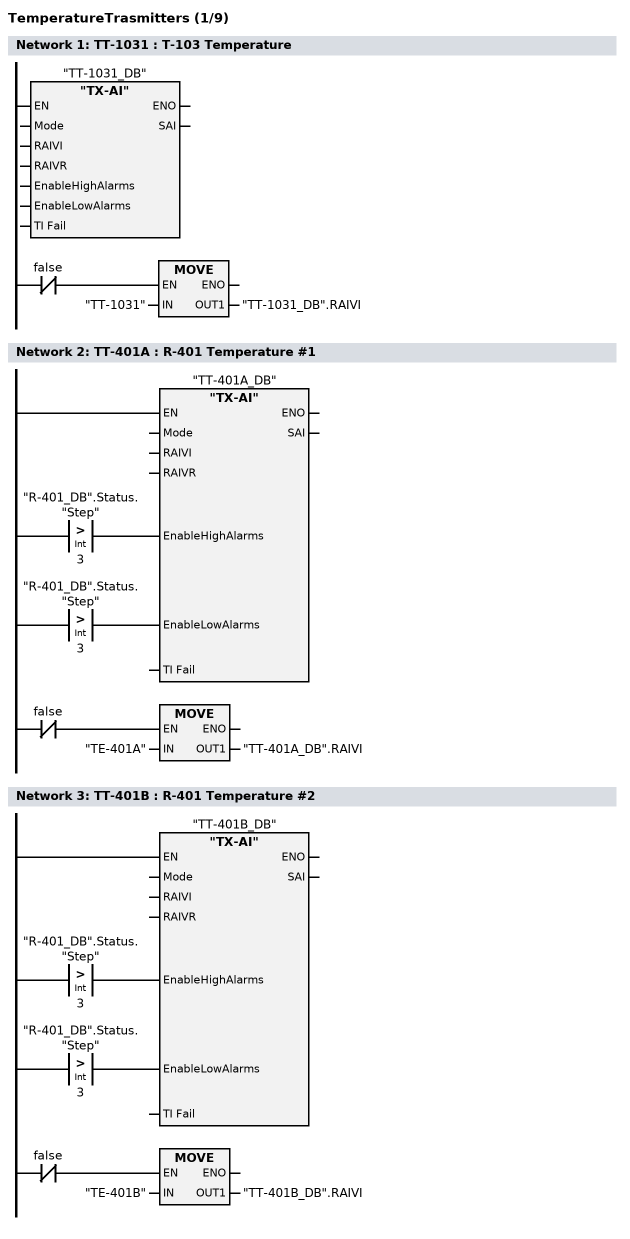
   RUNG wire#powerrail
      "TT-1031_DB"(Mode :=, RAIVI :=, RAIVR :=, EnableHighAlarms :=, EnableLowAlarms :=, "TI Fail" :=, SAI =>)
   END_RUNG
   RUNG wire#powerrail
      I_Contact( false )
      { S7_GenerateENO := "TRUE" } Move(in := "TT-1031", out1 => "TT-1031_DB".RAIVI)
   END_RUNG
   // the same network as SCL:
   "TT-1031_DB"();   // "TX-AI"
   IF NOT false THEN "TT-1031_DB".RAIVI := "TT-1031"; END_IF;
END_REGION

REGION Network 2: TT-401A : R-401 Temperature #1
   RUNG wire#powerrail
      "TT-401A_DB"(EnableHighAlarms := wire#w1, EnableLowAlarms := wire#w2, Mode :=, RAIVI :=, RAIVR :=, "TI Fail" :=, SAI =>)
   END_RUNG
   RUNG wire#powerrail
      { S7_Templates := "SrcType := Int" } GT_Contact(in1 := "R-401_DB".Status."Step", in2 := 3)
   END_RUNG wire#w1
   RUNG wire#powerrail
      { S7_Templates := "SrcType := Int" } GT_Contact(in1 := "R-401_DB".Status."Step", in2 := 3)
   END_RUNG wire#w2
   RUNG wire#powerrail
      I_Contact( false )
      { S7_GenerateENO := "TRUE" } Move(in := "TE-401A", out1 => "TT-401A_DB".RAIVI)
   END_RUNG
   // the same network as SCL:
   "TT-401A_DB"(EnableHighAlarms := "R-401_DB".Status."Step" > 3,   // "TX-AI"
                EnableLowAlarms := "R-401_DB".Status."Step" > 3);
   IF NOT false THEN "TT-401A_DB".RAIVI := "TE-401A"; END_IF;
END_REGION

REGION Network 3: TT-401B : R-401 Temperature #2
   RUNG wire#powerrail
      "TT-401B_DB"(EnableHighAlarms := wire#w1, EnableLowAlarms := wire#w2, Mode :=, RAIVI :=, RAIVR :=, "TI Fail" :=, SAI =>)
   END_RUNG
   RUNG wire#powerrail
      { S7_Templates := "SrcType := Int" } GT_Contact(in1 := "R-401_DB".Status."Step", in2 := 3)
   END_RUNG wire#w1
   RUNG wire#powerrail
      { S7_Templates := "SrcType := Int" } GT_Contact(in1 := "R-401_DB".Status."Step", in2 := 3)
   END_RUNG wire#w2
   RUNG wire#powerrail
      I_Contact( false )
      { S7_GenerateENO := "TRUE" } Move(in := "TE-401B", out1 => "TT-401B_DB".RAIVI)
   END_RUNG
   // the same network as SCL:
   "TT-401B_DB"(EnableHighAlarms := "R-401_DB".Status."Step" > 3,   // "TX-AI"
                EnableLowAlarms := "R-401_DB".Status."Step" > 3);
   IF NOT false THEN "TT-401B_DB".RAIVI := "TE-401B"; END_IF;
END_REGION

REGION Network 4: TT-401C : R-401 Temperature #3
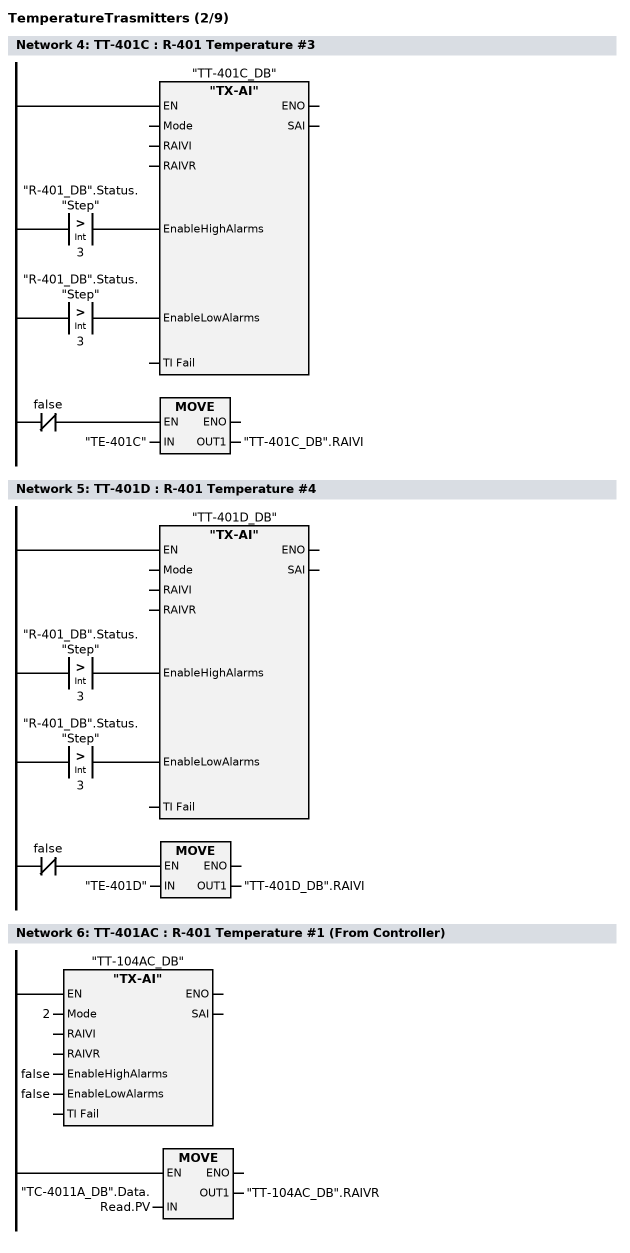
   RUNG wire#powerrail
      "TT-401C_DB"(EnableHighAlarms := wire#w1, EnableLowAlarms := wire#w2, Mode :=, RAIVI :=, RAIVR :=, "TI Fail" :=, SAI =>)
   END_RUNG
   RUNG wire#powerrail
      { S7_Templates := "SrcType := Int" } GT_Contact(in1 := "R-401_DB".Status."Step", in2 := 3)
   END_RUNG wire#w1
   RUNG wire#powerrail
      { S7_Templates := "SrcType := Int" } GT_Contact(in1 := "R-401_DB".Status."Step", in2 := 3)
   END_RUNG wire#w2
   RUNG wire#powerrail
      I_Contact( false )
      { S7_GenerateENO := "TRUE" } Move(in := "TE-401C", out1 => "TT-401C_DB".RAIVI)
   END_RUNG
   // the same network as SCL:
   "TT-401C_DB"(EnableHighAlarms := "R-401_DB".Status."Step" > 3,   // "TX-AI"
                EnableLowAlarms := "R-401_DB".Status."Step" > 3);
   IF NOT false THEN "TT-401C_DB".RAIVI := "TE-401C"; END_IF;
END_REGION

REGION Network 5: TT-401D : R-401 Temperature #4
   RUNG wire#powerrail
      "TT-401D_DB"(EnableHighAlarms := wire#w1, EnableLowAlarms := wire#w2, Mode :=, RAIVI :=, RAIVR :=, "TI Fail" :=, SAI =>)
   END_RUNG
   RUNG wire#powerrail
      { S7_Templates := "SrcType := Int" } GT_Contact(in1 := "R-401_DB".Status."Step", in2 := 3)
   END_RUNG wire#w1
   RUNG wire#powerrail
      { S7_Templates := "SrcType := Int" } GT_Contact(in1 := "R-401_DB".Status."Step", in2 := 3)
   END_RUNG wire#w2
   RUNG wire#powerrail
      I_Contact( false )
      { S7_GenerateENO := "TRUE" } Move(in := "TE-401D", out1 => "TT-401D_DB".RAIVI)
   END_RUNG
   // the same network as SCL:
   "TT-401D_DB"(EnableHighAlarms := "R-401_DB".Status."Step" > 3,   // "TX-AI"
                EnableLowAlarms := "R-401_DB".Status."Step" > 3);
   IF NOT false THEN "TT-401D_DB".RAIVI := "TE-401D"; END_IF;
END_REGION

REGION Network 6: TT-401AC : R-401 Temperature #1 (From Controller)
   RUNG wire#powerrail
      "TT-104AC_DB"(Mode := 2, RAIVI :=, RAIVR :=, EnableHighAlarms := false, EnableLowAlarms := false, "TI Fail" :=, SAI =>)
   END_RUNG
   RUNG wire#powerrail
      { S7_GenerateENO := "TRUE" } Move(in := "TC-4011A_DB".Data.Read.PV, out1 => "TT-104AC_DB".RAIVR)
   END_RUNG
   // the same network as SCL:
   "TT-104AC_DB"(Mode := 2, EnableHighAlarms := false, EnableLowAlarms := false);   // "TX-AI"
   "TT-104AC_DB".RAIVR := "TC-4011A_DB".Data.Read.PV;
END_REGION

REGION Network 7: TT-401BC : R-401 Temperature #2 (From Controller)
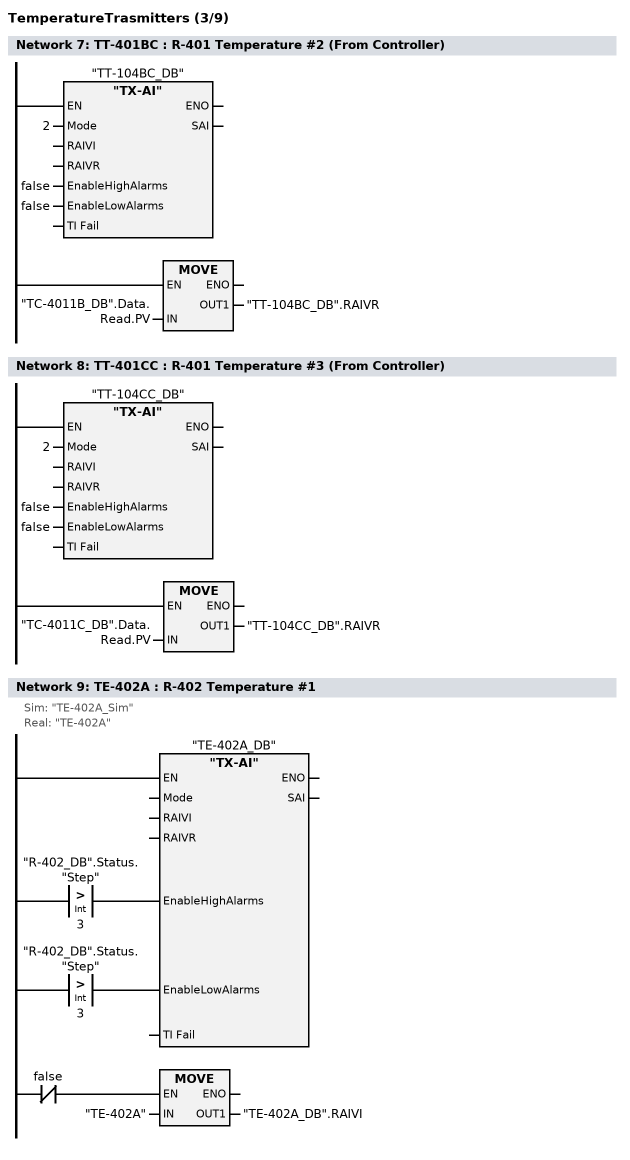
   RUNG wire#powerrail
      "TT-104BC_DB"(Mode := 2, RAIVI :=, RAIVR :=, EnableHighAlarms := false, EnableLowAlarms := false, "TI Fail" :=, SAI =>)
   END_RUNG
   RUNG wire#powerrail
      { S7_GenerateENO := "TRUE" } Move(in := "TC-4011B_DB".Data.Read.PV, out1 => "TT-104BC_DB".RAIVR)
   END_RUNG
   // the same network as SCL:
   "TT-104BC_DB"(Mode := 2, EnableHighAlarms := false, EnableLowAlarms := false);   // "TX-AI"
   "TT-104BC_DB".RAIVR := "TC-4011B_DB".Data.Read.PV;
END_REGION

REGION Network 8: TT-401CC : R-401 Temperature #3 (From Controller)
   RUNG wire#powerrail
      "TT-104CC_DB"(Mode := 2, RAIVI :=, RAIVR :=, EnableHighAlarms := false, EnableLowAlarms := false, "TI Fail" :=, SAI =>)
   END_RUNG
   RUNG wire#powerrail
      { S7_GenerateENO := "TRUE" } Move(in := "TC-4011C_DB".Data.Read.PV, out1 => "TT-104CC_DB".RAIVR)
   END_RUNG
   // the same network as SCL:
   "TT-104CC_DB"(Mode := 2, EnableHighAlarms := false, EnableLowAlarms := false);   // "TX-AI"
   "TT-104CC_DB".RAIVR := "TC-4011C_DB".Data.Read.PV;
END_REGION

REGION Network 9: TE-402A : R-402 Temperature #1
   // Sim: "TE-402A_Sim"
   // Real: "TE-402A"
   RUNG wire#powerrail
      "TE-402A_DB"(EnableHighAlarms := wire#w1, EnableLowAlarms := wire#w2, Mode :=, RAIVI :=, RAIVR :=, "TI Fail" :=, SAI =>)
   END_RUNG
   RUNG wire#powerrail
      { S7_Templates := "SrcType := Int" } GT_Contact(in1 := "R-402_DB".Status."Step", in2 := 3)
   END_RUNG wire#w1
   RUNG wire#powerrail
      { S7_Templates := "SrcType := Int" } GT_Contact(in1 := "R-402_DB".Status."Step", in2 := 3)
   END_RUNG wire#w2
   RUNG wire#powerrail
      I_Contact( false )
      { S7_GenerateENO := "TRUE" } Move(in := "TE-402A", out1 => "TE-402A_DB".RAIVI)
   END_RUNG
   // the same network as SCL:
   "TE-402A_DB"(EnableHighAlarms := "R-402_DB".Status."Step" > 3,   // "TX-AI"
                EnableLowAlarms := "R-402_DB".Status."Step" > 3);
   IF NOT false THEN "TE-402A_DB".RAIVI := "TE-402A"; END_IF;
END_REGION

REGION Network 10: TE-402B : R-402 Temperature #2
   // Sim: "TE-402B_Sim"
   // Real: "TE-402B"
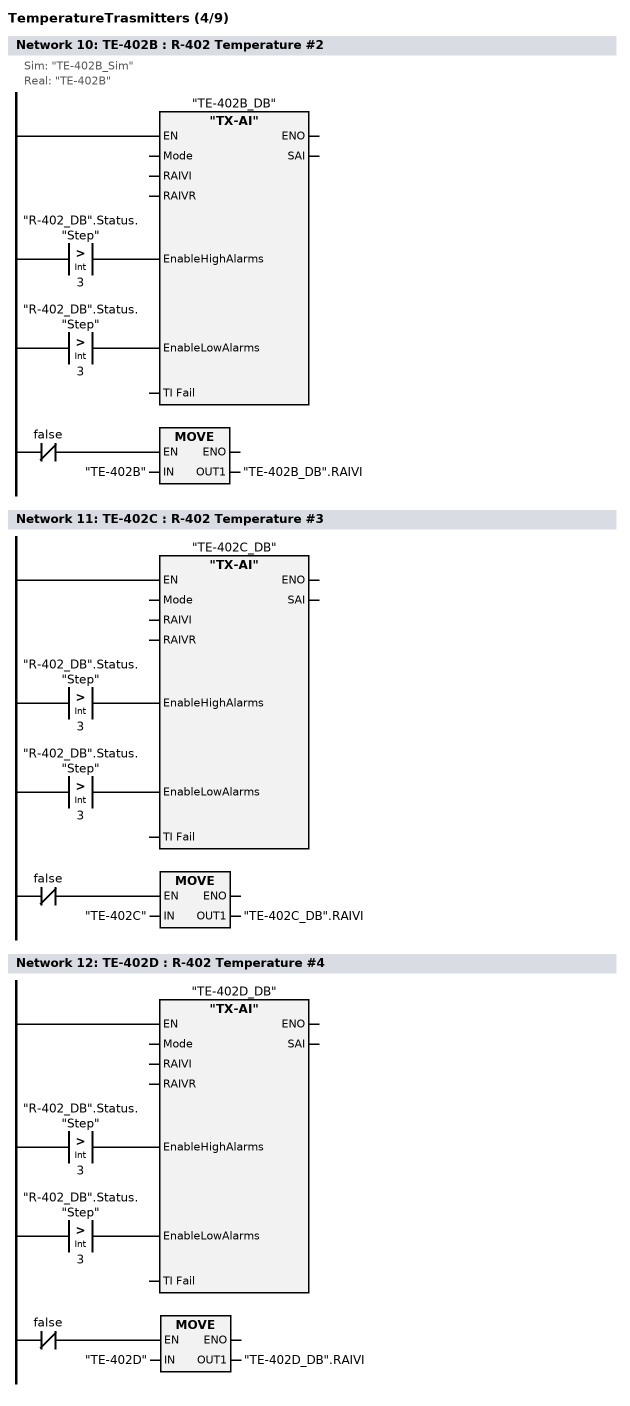
   RUNG wire#powerrail
      "TE-402B_DB"(EnableHighAlarms := wire#w1, EnableLowAlarms := wire#w2, Mode :=, RAIVI :=, RAIVR :=, "TI Fail" :=, SAI =>)
   END_RUNG
   RUNG wire#powerrail
      { S7_Templates := "SrcType := Int" } GT_Contact(in1 := "R-402_DB".Status."Step", in2 := 3)
   END_RUNG wire#w1
   RUNG wire#powerrail
      { S7_Templates := "SrcType := Int" } GT_Contact(in1 := "R-402_DB".Status."Step", in2 := 3)
   END_RUNG wire#w2
   RUNG wire#powerrail
      I_Contact( false )
      { S7_GenerateENO := "TRUE" } Move(in := "TE-402B", out1 => "TE-402B_DB".RAIVI)
   END_RUNG
   // the same network as SCL:
   "TE-402B_DB"(EnableHighAlarms := "R-402_DB".Status."Step" > 3,   // "TX-AI"
                EnableLowAlarms := "R-402_DB".Status."Step" > 3);
   IF NOT false THEN "TE-402B_DB".RAIVI := "TE-402B"; END_IF;
END_REGION

REGION Network 11: TE-402C : R-402 Temperature #3
   RUNG wire#powerrail
      "TE-402C_DB"(EnableHighAlarms := wire#w1, EnableLowAlarms := wire#w2, Mode :=, RAIVI :=, RAIVR :=, "TI Fail" :=, SAI =>)
   END_RUNG
   RUNG wire#powerrail
      { S7_Templates := "SrcType := Int" } GT_Contact(in1 := "R-402_DB".Status."Step", in2 := 3)
   END_RUNG wire#w1
   RUNG wire#powerrail
      { S7_Templates := "SrcType := Int" } GT_Contact(in1 := "R-402_DB".Status."Step", in2 := 3)
   END_RUNG wire#w2
   RUNG wire#powerrail
      I_Contact( false )
      { S7_GenerateENO := "TRUE" } Move(in := "TE-402C", out1 => "TE-402C_DB".RAIVI)
   END_RUNG
   // the same network as SCL:
   "TE-402C_DB"(EnableHighAlarms := "R-402_DB".Status."Step" > 3,   // "TX-AI"
                EnableLowAlarms := "R-402_DB".Status."Step" > 3);
   IF NOT false THEN "TE-402C_DB".RAIVI := "TE-402C"; END_IF;
END_REGION

REGION Network 12: TE-402D : R-402 Temperature #4
   RUNG wire#powerrail
      "TE-402D_DB"(EnableHighAlarms := wire#w1, EnableLowAlarms := wire#w2, Mode :=, RAIVI :=, RAIVR :=, "TI Fail" :=, SAI =>)
   END_RUNG
   RUNG wire#powerrail
      { S7_Templates := "SrcType := Int" } GT_Contact(in1 := "R-402_DB".Status."Step", in2 := 3)
   END_RUNG wire#w1
   RUNG wire#powerrail
      { S7_Templates := "SrcType := Int" } GT_Contact(in1 := "R-402_DB".Status."Step", in2 := 3)
   END_RUNG wire#w2
   RUNG wire#powerrail
      I_Contact( false )
      { S7_GenerateENO := "TRUE" } Move(in := "TE-402D", out1 => "TE-402D_DB".RAIVI)
   END_RUNG
   // the same network as SCL:
   "TE-402D_DB"(EnableHighAlarms := "R-402_DB".Status."Step" > 3,   // "TX-AI"
                EnableLowAlarms := "R-402_DB".Status."Step" > 3);
   IF NOT false THEN "TE-402D_DB".RAIVI := "TE-402D"; END_IF;
END_REGION

REGION Network 13: TE-402E : R-402 Temperature #5
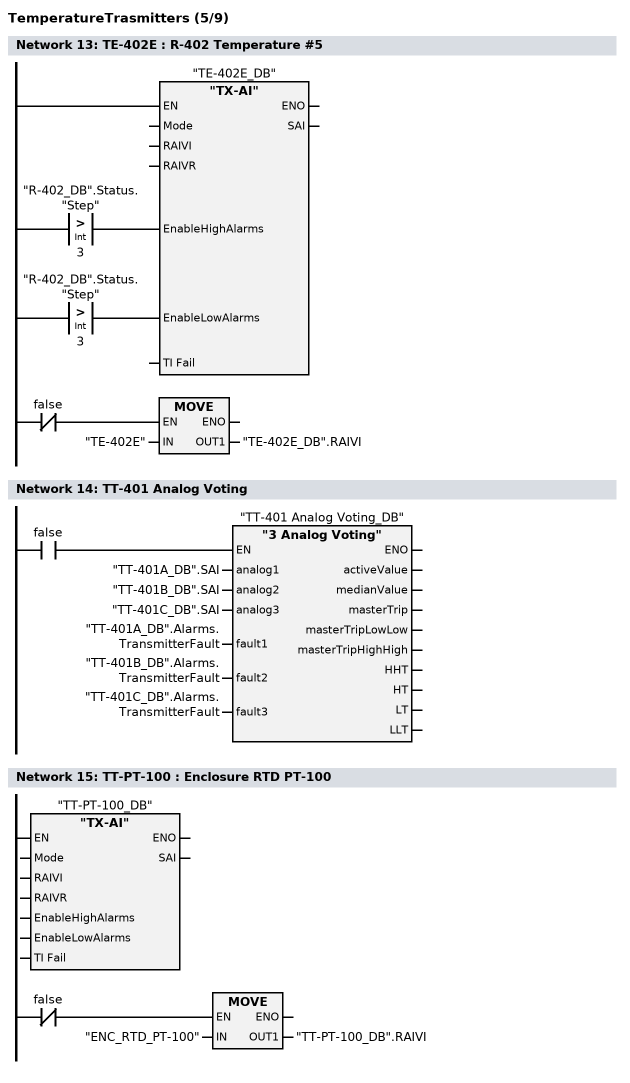
   RUNG wire#powerrail
      "TE-402E_DB"(EnableHighAlarms := wire#w1, EnableLowAlarms := wire#w2, Mode :=, RAIVI :=, RAIVR :=, "TI Fail" :=, SAI =>)
   END_RUNG
   RUNG wire#powerrail
      { S7_Templates := "SrcType := Int" } GT_Contact(in1 := "R-402_DB".Status."Step", in2 := 3)
   END_RUNG wire#w1
   RUNG wire#powerrail
      { S7_Templates := "SrcType := Int" } GT_Contact(in1 := "R-402_DB".Status."Step", in2 := 3)
   END_RUNG wire#w2
   RUNG wire#powerrail
      I_Contact( false )
      { S7_GenerateENO := "TRUE" } Move(in := "TE-402E", out1 => "TE-402E_DB".RAIVI)
   END_RUNG
   // the same network as SCL:
   "TE-402E_DB"(EnableHighAlarms := "R-402_DB".Status."Step" > 3,   // "TX-AI"
                EnableLowAlarms := "R-402_DB".Status."Step" > 3);
   IF NOT false THEN "TE-402E_DB".RAIVI := "TE-402E"; END_IF;
END_REGION

REGION Network 14: TT-401 Analog Voting
   RUNG wire#powerrail
      Contact( false )
      "TT-401 Analog Voting_DB"(analog1 := "TT-401A_DB".SAI, analog2 := "TT-401B_DB".SAI, analog3 := "TT-401C_DB".SAI, fault1 := "TT-401A_DB".Alarms.TransmitterFault, fault2 := "TT-401B_DB".Alarms.TransmitterFault, fault3 := "TT-401C_DB".Alarms.TransmitterFault, activeValue =>, medianValue =>, masterTrip =>, masterTripLowLow =>, masterTripHighHigh =>, HHT =>, HT =>, LT =>, LLT =>)
   END_RUNG
   // the same network as SCL:
   IF false THEN
       "TT-401 Analog Voting_DB"(analog1 := "TT-401A_DB".SAI,   // "3 Analog Voting"
                               analog2 := "TT-401B_DB".SAI,
                               analog3 := "TT-401C_DB".SAI,
                               fault1 := "TT-401A_DB".Alarms.TransmitterFault,
                               fault2 := "TT-401B_DB".Alarms.TransmitterFault,
                               fault3 := "TT-401C_DB".Alarms.TransmitterFault);
   END_IF;
END_REGION

REGION Network 15: TT-PT-100 : Enclosure RTD PT-100
   RUNG wire#powerrail
      "TT-PT-100_DB"(Mode :=, RAIVI :=, RAIVR :=, EnableHighAlarms :=, EnableLowAlarms :=, "TI Fail" :=, SAI =>)
   END_RUNG
   RUNG wire#powerrail
      I_Contact( false )
      { S7_GenerateENO := "TRUE" } Move(in := "ENC_RTD_PT-100", out1 => "TT-PT-100_DB".RAIVI)
   END_RUNG
   // the same network as SCL:
   "TT-PT-100_DB"();   // "TX-AI"
   IF NOT false THEN "TT-PT-100_DB".RAIVI := "ENC_RTD_PT-100"; END_IF;
END_REGION

REGION Network 16: TT-2012 : R-201 Temperature #2
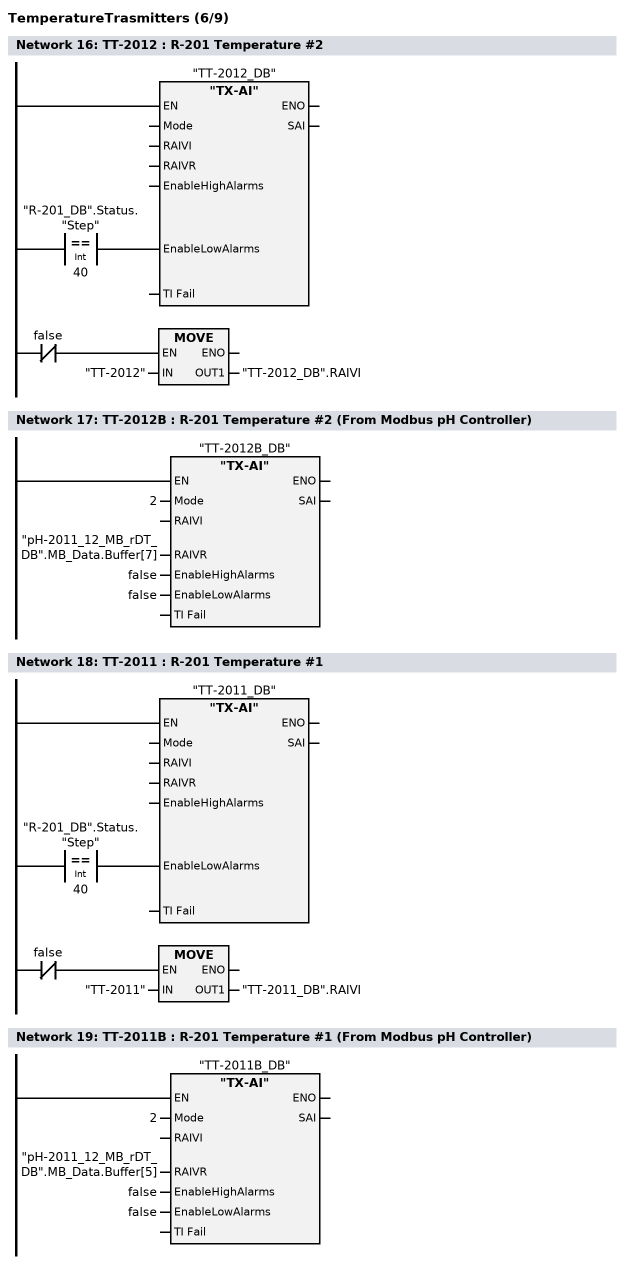
   RUNG wire#powerrail
      "TT-2012_DB"(EnableLowAlarms := wire#w1, Mode :=, RAIVI :=, RAIVR :=, EnableHighAlarms :=, "TI Fail" :=, SAI =>)
   END_RUNG
   RUNG wire#powerrail
      { S7_Templates := "SrcType := Int" } EQ_Contact(in1 := "R-201_DB".Status."Step", in2 := 40)
   END_RUNG wire#w1
   RUNG wire#powerrail
      I_Contact( false )
      { S7_GenerateENO := "TRUE" } Move(in := "TT-2012", out1 => "TT-2012_DB".RAIVI)
   END_RUNG
   // the same network as SCL:
   "TT-2012_DB"(EnableLowAlarms := "R-201_DB".Status."Step" = 40);   // "TX-AI"
   IF NOT false THEN "TT-2012_DB".RAIVI := "TT-2012"; END_IF;
END_REGION

REGION Network 17: TT-2012B : R-201 Temperature #2 (From Modbus pH Controller)
   RUNG wire#powerrail
      "TT-2012B_DB"(Mode := 2, RAIVI :=, RAIVR := "pH-2011_12_MB_rDT_DB".MB_Data.Buffer[7], EnableHighAlarms := false, EnableLowAlarms := false, "TI Fail" :=, SAI =>)
   END_RUNG
   // the same network as SCL:
   "TT-2012B_DB"(Mode := 2,   // "TX-AI"
                 RAIVR := "pH-2011_12_MB_rDT_DB".MB_Data.Buffer[7],
                 EnableHighAlarms := false,
                 EnableLowAlarms := false);
END_REGION

REGION Network 18: TT-2011 : R-201 Temperature #1
   RUNG wire#powerrail
      "TT-2011_DB"(EnableLowAlarms := wire#w1, Mode :=, RAIVI :=, RAIVR :=, EnableHighAlarms :=, "TI Fail" :=, SAI =>)
   END_RUNG
   RUNG wire#powerrail
      { S7_Templates := "SrcType := Int" } EQ_Contact(in1 := "R-201_DB".Status."Step", in2 := 40)
   END_RUNG wire#w1
   RUNG wire#powerrail
      I_Contact( false )
      { S7_GenerateENO := "TRUE" } Move(in := "TT-2011", out1 => "TT-2011_DB".RAIVI)
   END_RUNG
   // the same network as SCL:
   "TT-2011_DB"(EnableLowAlarms := "R-201_DB".Status."Step" = 40);   // "TX-AI"
   IF NOT false THEN "TT-2011_DB".RAIVI := "TT-2011"; END_IF;
END_REGION

REGION Network 19: TT-2011B : R-201 Temperature #1 (From Modbus pH Controller)
   RUNG wire#powerrail
      "TT-2011B_DB"(Mode := 2, RAIVI :=, RAIVR := "pH-2011_12_MB_rDT_DB".MB_Data.Buffer[5], EnableHighAlarms := false, EnableLowAlarms := false, "TI Fail" :=, SAI =>)
   END_RUNG
   // the same network as SCL:
   "TT-2011B_DB"(Mode := 2,   // "TX-AI"
                 RAIVR := "pH-2011_12_MB_rDT_DB".MB_Data.Buffer[5],
                 EnableHighAlarms := false,
                 EnableLowAlarms := false);
END_REGION

REGION Network 20: R-201 Temperature Average
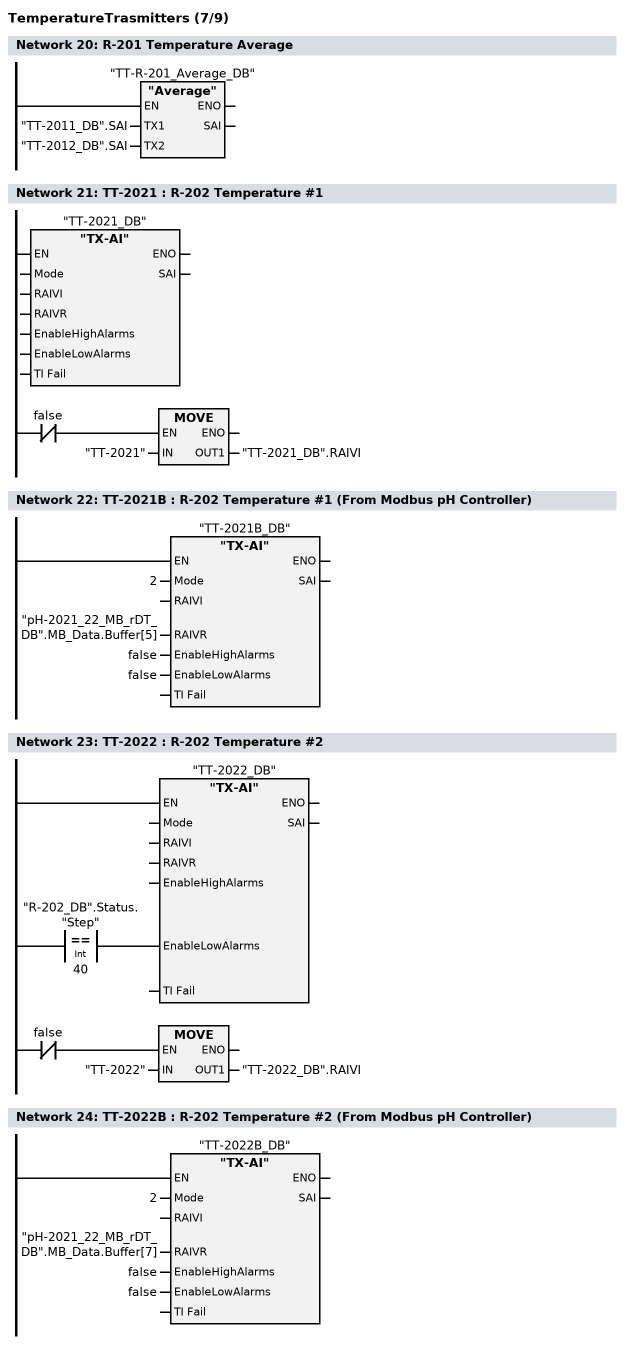
   RUNG wire#powerrail
      "TT-R-201_Average_DB"(TX1 := "TT-2011_DB".SAI, TX2 := "TT-2012_DB".SAI, SAI =>)
   END_RUNG
   // the same network as SCL:
   "TT-R-201_Average_DB"(TX1 := "TT-2011_DB".SAI, TX2 := "TT-2012_DB".SAI);   // "Average"
END_REGION

REGION Network 21: TT-2021 : R-202 Temperature #1
   RUNG wire#powerrail
      "TT-2021_DB"(Mode :=, RAIVI :=, RAIVR :=, EnableHighAlarms :=, EnableLowAlarms :=, "TI Fail" :=, SAI =>)
   END_RUNG
   RUNG wire#powerrail
      I_Contact( false )
      { S7_GenerateENO := "TRUE" } Move(in := "TT-2021", out1 => "TT-2021_DB".RAIVI)
   END_RUNG
   // the same network as SCL:
   "TT-2021_DB"();   // "TX-AI"
   IF NOT false THEN "TT-2021_DB".RAIVI := "TT-2021"; END_IF;
END_REGION

REGION Network 22: TT-2021B : R-202 Temperature #1 (From Modbus pH Controller)
   RUNG wire#powerrail
      "TT-2021B_DB"(Mode := 2, RAIVI :=, RAIVR := "pH-2021_22_MB_rDT_DB".MB_Data.Buffer[5], EnableHighAlarms := false, EnableLowAlarms := false, "TI Fail" :=, SAI =>)
   END_RUNG
   // the same network as SCL:
   "TT-2021B_DB"(Mode := 2,   // "TX-AI"
                 RAIVR := "pH-2021_22_MB_rDT_DB".MB_Data.Buffer[5],
                 EnableHighAlarms := false,
                 EnableLowAlarms := false);
END_REGION

REGION Network 23: TT-2022 : R-202 Temperature #2
   RUNG wire#powerrail
      "TT-2022_DB"(EnableLowAlarms := wire#w1, Mode :=, RAIVI :=, RAIVR :=, EnableHighAlarms :=, "TI Fail" :=, SAI =>)
   END_RUNG
   RUNG wire#powerrail
      { S7_Templates := "SrcType := Int" } EQ_Contact(in1 := "R-202_DB".Status."Step", in2 := 40)
   END_RUNG wire#w1
   RUNG wire#powerrail
      I_Contact( false )
      { S7_GenerateENO := "TRUE" } Move(in := "TT-2022", out1 => "TT-2022_DB".RAIVI)
   END_RUNG
   // the same network as SCL:
   "TT-2022_DB"(EnableLowAlarms := "R-202_DB".Status."Step" = 40);   // "TX-AI"
   IF NOT false THEN "TT-2022_DB".RAIVI := "TT-2022"; END_IF;
END_REGION

REGION Network 24: TT-2022B : R-202 Temperature #2 (From Modbus pH Controller)
   RUNG wire#powerrail
      "TT-2022B_DB"(Mode := 2, RAIVI :=, RAIVR := "pH-2021_22_MB_rDT_DB".MB_Data.Buffer[7], EnableHighAlarms := false, EnableLowAlarms := false, "TI Fail" :=, SAI =>)
   END_RUNG
   // the same network as SCL:
   "TT-2022B_DB"(Mode := 2,   // "TX-AI"
                 RAIVR := "pH-2021_22_MB_rDT_DB".MB_Data.Buffer[7],
                 EnableHighAlarms := false,
                 EnableLowAlarms := false);
END_REGION

REGION Network 25: R-202 Temperature Average
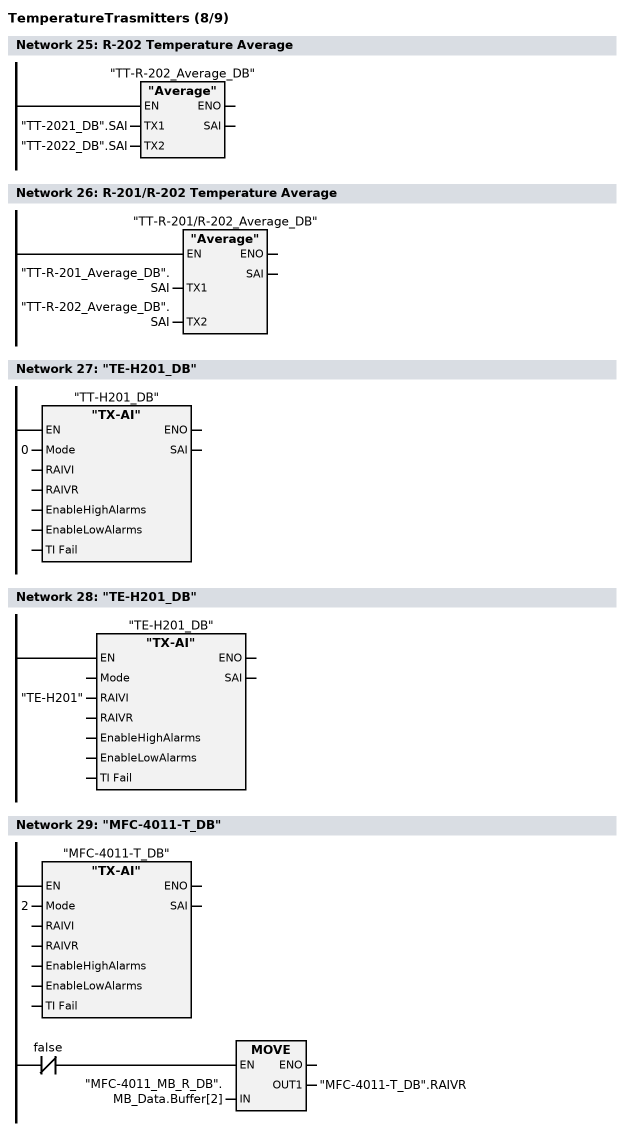
   RUNG wire#powerrail
      "TT-R-202_Average_DB"(TX1 := "TT-2021_DB".SAI, TX2 := "TT-2022_DB".SAI, SAI =>)
   END_RUNG
   // the same network as SCL:
   "TT-R-202_Average_DB"(TX1 := "TT-2021_DB".SAI, TX2 := "TT-2022_DB".SAI);   // "Average"
END_REGION

REGION Network 26: R-201/R-202 Temperature Average
   RUNG wire#powerrail
      "TT-R-201/R-202_Average_DB"(TX1 := "TT-R-201_Average_DB".SAI, TX2 := "TT-R-202_Average_DB".SAI, SAI =>)
   END_RUNG
   // the same network as SCL:
   "TT-R-201/R-202_Average_DB"(TX1 := "TT-R-201_Average_DB".SAI, TX2 := "TT-R-202_Average_DB".SAI);   // "Average"
END_REGION

REGION Network 27: "TE-H201_DB"
   RUNG wire#powerrail
      "TT-H201_DB"(Mode := 0, RAIVI :=, RAIVR :=, EnableHighAlarms :=, EnableLowAlarms :=, "TI Fail" :=, SAI =>)
   END_RUNG
   // the same network as SCL:
   "TT-H201_DB"(Mode := 0);   // "TX-AI"
END_REGION

REGION Network 28: "TE-H201_DB"
   RUNG wire#powerrail
      "TE-H201_DB"(Mode :=, RAIVI := "TE-H201", RAIVR :=, EnableHighAlarms :=, EnableLowAlarms :=, "TI Fail" :=, SAI =>)
   END_RUNG
   // the same network as SCL:
   "TE-H201_DB"(RAIVI := "TE-H201");   // "TX-AI"
END_REGION

REGION Network 29: "MFC-4011-T_DB"
   RUNG wire#powerrail
      "MFC-4011-T_DB"(Mode := 2, RAIVI :=, RAIVR :=, EnableHighAlarms :=, EnableLowAlarms :=, "TI Fail" :=, SAI =>)
   END_RUNG
   RUNG wire#powerrail
      I_Contact( false )
      { S7_GenerateENO := "TRUE" } Move(in := "MFC-4011_MB_R_DB".MB_Data.Buffer[2], out1 => "MFC-4011-T_DB".RAIVR)
   END_RUNG
   // the same network as SCL:
   "MFC-4011-T_DB"(Mode := 2);   // "TX-AI"
   IF NOT false THEN "MFC-4011-T_DB".RAIVR := "MFC-4011_MB_R_DB".MB_Data.Buffer[2]; END_IF;
END_REGION

REGION Network 30: "MFC-4012-T_DB"
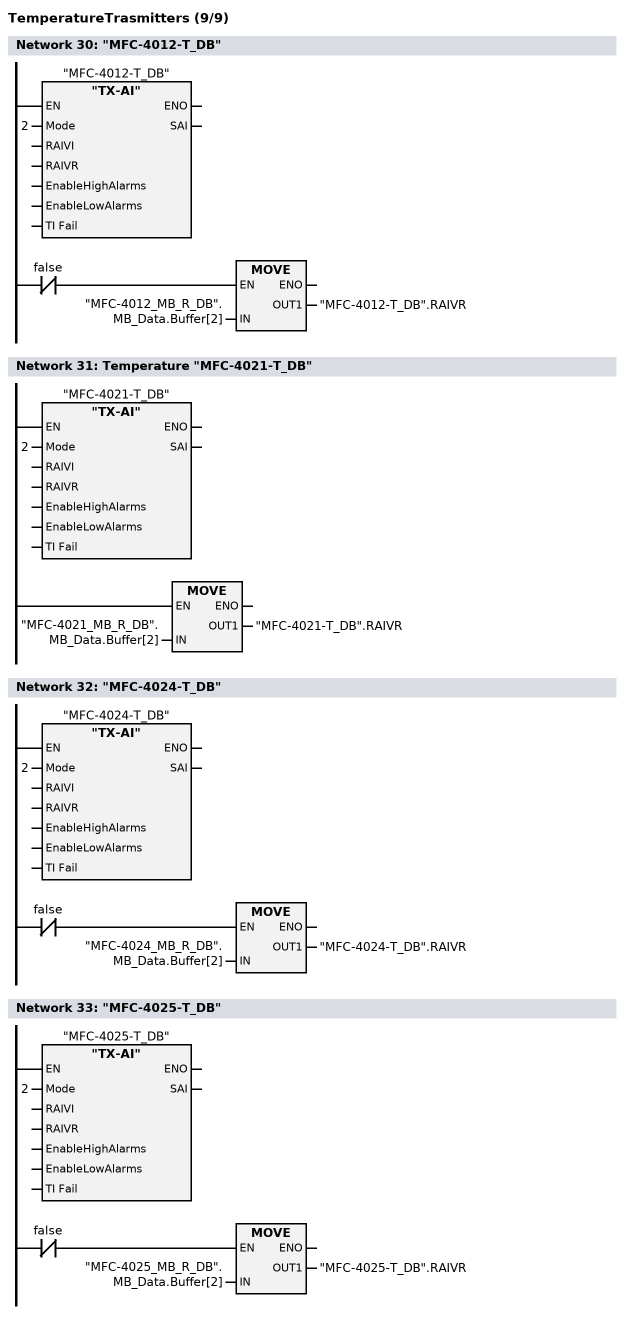
   RUNG wire#powerrail
      "MFC-4012-T_DB"(Mode := 2, RAIVI :=, RAIVR :=, EnableHighAlarms :=, EnableLowAlarms :=, "TI Fail" :=, SAI =>)
   END_RUNG
   RUNG wire#powerrail
      I_Contact( false )
      { S7_GenerateENO := "TRUE" } Move(in := "MFC-4012_MB_R_DB".MB_Data.Buffer[2], out1 => "MFC-4012-T_DB".RAIVR)
   END_RUNG
   // the same network as SCL:
   "MFC-4012-T_DB"(Mode := 2);   // "TX-AI"
   IF NOT false THEN "MFC-4012-T_DB".RAIVR := "MFC-4012_MB_R_DB".MB_Data.Buffer[2]; END_IF;
END_REGION

REGION Network 31: Temperature "MFC-4021-T_DB"
   RUNG wire#powerrail
      "MFC-4021-T_DB"(Mode := 2, RAIVI :=, RAIVR :=, EnableHighAlarms :=, EnableLowAlarms :=, "TI Fail" :=, SAI =>)
   END_RUNG
   RUNG wire#powerrail
      { S7_GenerateENO := "TRUE" } Move(in := "MFC-4021_MB_R_DB".MB_Data.Buffer[2], out1 => "MFC-4021-T_DB".RAIVR)
   END_RUNG
   // the same network as SCL:
   "MFC-4021-T_DB"(Mode := 2);   // "TX-AI"
   "MFC-4021-T_DB".RAIVR := "MFC-4021_MB_R_DB".MB_Data.Buffer[2];
END_REGION
